VERSION : 1.2
// clk_pulse uses the internal sps time to generate a clock with programmable period time.
// the period time is defined for 10ms .. 65s.
// pulse generation is continuous if N = 0 and for n pulses otherwise.
// the first cycle after start is a clk pulse and then depending on the programmed period time a delay.
// every pulse is only valid for one cycle so that a edge trigger is not necessary
// clk_prg depending on the accuracy of the system clock.
// 
// uses: T_PLC_MS [FC64]
//       STIME [FB64],IDB_STIME [DB64]
   VAR_INPUT
      PT : Time;
      N : Int;
      RST : Bool;
   END_VAR
   VAR_OUTPUT
      Q : Bool;
      CNT : Int;
      RUN : Bool;
   END_VAR
   VAR
      tx : DWord;
      tn : DWord;
      init : Bool;
   END_VAR
   VAR_TEMP
      TOP_SI : Struct
         EV_CLASS : Byte;
         EV_NUM : Byte;
         PRIORITY : Byte;
         NUM : Byte;
         TYP2_3 : Byte;
         TYP1 : Byte;
         ZI1 : Word;
         ZI2_3 : DWord;
      END_STRUCT;
      START_UP_SI : Struct
         EV_CLASS : Byte;
         EV_NUM : Byte;
         PRIORITY : Byte;
         NUM : Byte;
         TYP2_3 : Byte;
         TYP1 : Byte;
         ZI1 : Word;
         ZI2_3 : DWord;
      END_STRUCT;
      ERR : Int;
   END_VAR
BEGIN


   (* read actual startup info *)
   (* OB1_SCAN_1  BYTE  -  B#16#01: Abschluss des Neustarts (Warmstarts)
                        -  B#16#02: Abschluss des Wiederanlaufs
                        -  B#16#03: Abschluss des freien Zyklus
                        -  B#16#04: Abschluss des Kaltstarts
                        -  B#16#05: Erster OB 1-Zyklus der neuen Master-CPU nach 
                                    Master-Reserve-Umschaltung und STOP des 
                                    bisherigen Masters *)

     #ERR := RD_SINFO (TOP_SI => #TOP_SI, START_UP_SI => #START_UP_SI);

   (* detect system startup *)
     IF #TOP_SI.EV_NUM = 1 OR #TOP_SI.EV_NUM = 2 OR #TOP_SI.EV_NUM = 4 THEN 
       #init := FALSE;
     END_IF;

     #tx := "T_PLC_MS"();   (* read system *)
     #Q := FALSE;       (* reset Q we generate pulses only for one cycle *)
     #RUN := #CNT < #N;

     IF NOT #init OR #RST THEN
       #init := TRUE;
       #CNT := 0;
       #tn := DINT_TO_DWORD(DWORD_TO_DINT(#tx) - T_CONV(#PT));
       #RUN := FALSE;
     ELSIF (#CNT < #N OR #N = 0) AND DWORD_TO_DINT(#tx) - DWORD_TO_DINT(#tn) >= T_CONV(#PT) THEN    (* generate a pulse *)
       #CNT := #CNT + 1;
       #Q := TRUE;
       #tn := DINT_TO_DWORD(DWORD_TO_DINT(#tn) + T_CONV(#PT));
     END_IF;


   (* revision history
   hm    4. aug 2006   rev 1.0
     original version

   hm    17. sep 2007  rev 1.1
     replaced time() with T_PLC_S() for compatblity reasons

   hm    16. feb. 2011 rev 1.2
     fixed an error when timer overflows 
   *)
END_FUNCTION_BLOCK

FUNCTION_BLOCK "D_TRIG"   // FB54, SCL
TITLE = D_TRIG
{ S7_Optimized_Access := 'FALSE' }
AUTHOR : hugo
FAMILY : GENERAT
NAME : D_TRIG
VERSION : 1.1
// this block is similar to the IEC Standard R_trig and F_trig but it monitors a DWORD, WORD or Byte Variable instead and generated an Output Pulse for one cycle only when the input has changed.
// an additional output x (Dword) will state the chage of the input.
// Example: the input has chaged from 0001 to 0010 then the output x will be 2.
   VAR_INPUT
      in : DWord;
   END_VAR
   VAR_OUTPUT
      Q : Bool;
      X : DWord;
   END_VAR
   VAR
      last_in : DWord;
   END_VAR
BEGIN


     #Q := #in <> #last_in;
     #X := DINT_TO_DWORD(DWORD_TO_DINT(#in) - DWORD_TO_DINT(#last_in));
     #last_in := #in;


   (* revision history

   hm  4.09.2007   rev 1.0
     original version released

   hm  19. feb. 2008 rev 1.1
     performance improvement
   *)
END_FUNCTION_BLOCK

FUNCTION_BLOCK "GEN_BIT"   // FB55, SCL
TITLE = GEN_BIT
{ S7_Optimized_Access := 'FALSE' }
AUTHOR : hugo
FAMILY : GENERAT
NAME : GEN_BIT
VERSION : 1.2
// gen_bit is 4 bit sequencial pattern generator with 4 DWORD inputs and 4 serial outputs.
// with the first clock pulse after a reset or after power on, bit 0 of the input DWORDS IN is present on the Outputs Q and the next clock cycle shifts to Bit 1 and so on.
// the input steps defines how many bits of the input dwords will be shifted to the outputs. the sequence can be repetive when rep = 0 or any amount of repetitions can be defined with input rep.
   VAR_INPUT
      in0 : DWord;
      in1 : DWord;
      in2 : DWord;
      in3 : DWord;
      clk : Bool;
      steps : Int;
      rep : Int;
      rst : Bool;
   END_VAR
   VAR_OUTPUT
      Q0 : Bool;
      Q1 : Bool;
      Q2 : Bool;
      Q3 : Bool;
      cnt : Int;
      run : Bool;
   END_VAR
   VAR
      r0 : DWord;
      tr0 AT r0 : Array[0..31] of Bool;
      r1 : DWord;
      tr1 AT r1 : Array[0..31] of Bool;
      r2 : DWord;
      tr2 AT r2 : Array[0..31] of Bool;
      r3 : DWord;
      tr3 AT r3 : Array[0..31] of Bool;
      rx : Int := 1;
   END_VAR
BEGIN


   (* check if number of runs is finished or rep = 0 which means continuous *)
   IF #clk AND NOT #rst THEN
       #run := (#rep = 0) OR (#rx <= #rep);
       IF #run THEN
           (* check for step counter reached and reset to 0 if cnt = steps *)
           IF #cnt = #steps THEN
               #cnt := 0;
           END_IF;

           (* when cnt = 0 then reload the inputs into the registers *)
           IF #cnt = 0 THEN
               #r0 := #in0;
               #r1 := #in1;
               #r2 := #in2;
               #r3 := #in3;
           END_IF;

           (* when cnt < steps, shift the lowest bits to the outputs *)
           IF (#cnt < #steps) THEN
               #Q0 := #tr0[24];
               #Q1 := #tr1[24];
               #Q2 := #tr2[24];
               #Q3 := #tr3[24];
               #r0 := SHR(IN:=#r0,N:=1);
               #r1 := SHR(IN:=#r1,N:=1);
               #r2 := SHR(IN:=#r2,N:=1);
               #r3 := SHR(IN:=#r3,N:=1);
           END_IF;

           (* increment the step counter *)
           #cnt := #cnt +1;
           IF (#cnt = #steps) AND (#rep <> 0) THEN #rx := #rx +1; END_IF;
           IF (#rx > #rep) AND (#rep <> 0) THEN #run := FALSE; END_IF;
       END_IF;
   ELSE
       IF #rst THEN
           #run := FALSE;
           #Q0 := FALSE;
           #Q1 := FALSE;
           #Q2 := FALSE;
           #Q3 := FALSE;
           #r0 := 0;
           #r1 := 0;
           #r2 := 0;
           #r3 := 0;
           #cnt := 0;
           #rx := 1;
       END_IF;
   END_IF;


   (* revision histroy
   hm  4 aug 2006  rev 1.0
       original version

   hm 15. oct. 2008    rev 1.1
       improved performance

   hm  14. mar. 2009   rev 1.2
       removed double assignments

   *)
END_FUNCTION_BLOCK

FUNCTION_BLOCK "GEN_SQ"   // FB56, SCL
TITLE = GEN_SQ
{ S7_Optimized_Access := 'FALSE' }
AUTHOR : hugo
FAMILY : GENERAT
NAME : GEN_SQ
VERSION : 1.3
// gen_sq generates square wave signal with programmable period time.
// 
// uses: T_PLC_MS [FC64]
//       STIME [FB64],IDB_STIME [DB64]
   VAR_INPUT
      PT : Time;
   END_VAR
   VAR_OUTPUT
      Q : Bool;
   END_VAR
   VAR
      tn : Time;
      tx : Time;
      init : Bool;
   END_VAR
   VAR_TEMP
      TOP_SI : Struct
         EV_CLASS : Byte;
         EV_NUM : Byte;
         PRIORITY : Byte;
         NUM : Byte;
         TYP2_3 : Byte;
         TYP1 : Byte;
         ZI1 : Word;
         ZI2_3 : DWord;
      END_STRUCT;
      START_UP_SI : Struct
         EV_CLASS : Byte;
         EV_NUM : Byte;
         PRIORITY : Byte;
         NUM : Byte;
         TYP2_3 : Byte;
         TYP1 : Byte;
         ZI1 : Word;
         ZI2_3 : DWord;
      END_STRUCT;
      ERR : Int;
   END_VAR
BEGIN


     (* read actual startup info *)
     (* OB1_SCAN_1  BYTE  -  B#16#01: Abschluss des Neustarts (Warmstarts)
                          -  B#16#02: Abschluss des Wiederanlaufs
                          -  B#16#03: Abschluss des freien Zyklus
                          -  B#16#04: Abschluss des Kaltstarts
                          -  B#16#05: Erster OB 1-Zyklus der neuen Master-CPU nach 
                                      Master-Reserve-Umschaltung und STOP des 
                                      bisherigen Masters *)

     #ERR := RD_SINFO (TOP_SI => #TOP_SI, START_UP_SI => #START_UP_SI);

     (* read system time *)
     #tx := T_CONV(DWORD_TO_DINT("T_PLC_MS"()));

     (* reset last_time on system startup *)
     IF #TOP_SI.EV_NUM = 1 OR #TOP_SI.EV_NUM = 2 OR #TOP_SI.EV_NUM = 4 THEN 
       #init := FALSE;
     END_IF;

     IF NOT #init THEN
       #init := TRUE;
       #tn := #tx;
       #Q := TRUE;
     ELSIF #tx - #tn >= T_CONV(DWORD_TO_DINT(SHR(IN:=DINT_TO_DWORD(T_CONV(#PT)),N:=1))) THEN
       #Q := NOT #Q;
       #tn := #tn + T_CONV(DWORD_TO_DINT(SHR(IN:=DINT_TO_DWORD(T_CONV(#PT)),N:=1)));
     END_IF;


   (* revision history
   hm  4. aug 2006 rev 1.0
     original version

   hm  17. sep 2007  rev 1.1
     replaced time() with T_PLC_MS() for compatibility reasons

   hm  18. jul. 2009 rev 1.2
     improved accuracy

   hm  16. feb 2011  rev 1.3
     corrected an error with timer overflow 
   *)
END_FUNCTION_BLOCK

FUNCTION_BLOCK "SCHEDULER"   // FB57, SCL
TITLE = SCHEDULER
{ S7_Optimized_Access := 'FALSE' }
AUTHOR : hugo
FAMILY : GENERAT
NAME : SCHED
VERSION : 1.1
// SCHEDULER is used to call programs or function blocks at specific intervals.
// T0..T3 defines the interval times.
// 
// uses: T_PLC_MS [FC64]
//       STIME [FB64],IDB_STIME [DB64]
   VAR_INPUT
      E0 : Bool;
      E1 : Bool;
      E2 : Bool;
      E3 : Bool;
      T_0 : Time;
      T_1 : Time;
      T_2 : Time;
      T_3 : Time;
   END_VAR
   VAR_OUTPUT
      Q0 : Bool;
      Q1 : Bool;
      Q2 : Bool;
      Q3 : Bool;
   END_VAR
   VAR
      init : Bool;
      s0 : Time;
      s1 : Time;
      s2 : Time;
      s3 : Time;
      tx : Time;
      c : Int;
   END_VAR
BEGIN


   (* read system_time *)
   #tx := T_CONV(DWORD_TO_DINT("T_PLC_MS"()));

   IF NOT #init THEN
       #init := TRUE;
       #s0 := #tx - #T_0;
       #s1 := #tx - #T_1;
       #s2 := #tx - #T_2;
       #s3 := #tx - #T_3;
   END_IF;

   #Q0 := FALSE;
   #Q1 := FALSE;
   #Q2 := FALSE;
   #Q3 := FALSE;

   CASE #c OF
       0:  IF #tx - #s0 >= #T_0 THEN
               #Q0 := #E0;
               #s0 := #tx;
           END_IF;
           #c := 1;
       1:  IF #tx - #s1 >= #T_1 THEN
               #Q1 := #E1;
               #s1 := #tx;
           END_IF;
           #c := 2;
       2:  IF #tx - #s2 >= #T_2 THEN
               #Q2 := #E2;
               #s2 := #tx;
           END_IF;
           #c := 3;
       3:  IF #tx - #s3 >= #T_3 THEN
               #Q3 := #E3;
               #s3 := #tx;
           END_IF;
           #c := 0;
   END_CASE;


   (* revision history

   hm 28. sep. 2008    rev 1.0
       original version

   hm  14. mar. 2009   rev 1.1
       removed double assignments

   *)
END_FUNCTION_BLOCK

FUNCTION_BLOCK "SCHEDULER_2"   // FB58, SCL
TITLE = SCHEDULER_2
{ S7_Optimized_Access := 'FALSE' }
AUTHOR : hugo
FAMILY : GENERAT
NAME : SCHED2
VERSION : 1.0
// SCHEDULER_2 is used to call programs or function blocks at specific cycles.
// C0..C3 defines after how many cycles the output becomes active.
// O0..O3 defines a cycle offset at startup.
   VAR_INPUT
      E0 : Bool;
      E1 : Bool;
      E2 : Bool;
      E3 : Bool;
      C0 : Int;
      C1 : Int;
      C2 : Int;
      C3 : Int;
      O0 : Int;
      O1 : Int;
      O2 : Int;
      O3 : Int;
   END_VAR
   VAR_OUTPUT
      Q0 : Bool;
      Q1 : Bool;
      Q2 : Bool;
      Q3 : Bool;
   END_VAR
   VAR
      sx : Int;
   END_VAR
BEGIN


   #Q0 := #E0 AND (#sx MOD #C0 - #O0 = 0);
   #Q1 := #E1 AND (#sx MOD #C1 - #O1 = 0);
   #Q2 := #E2 AND (#sx MOD #C2 - #O2 = 0);
   #Q3 := #E3 AND (#sx MOD #C3 - #O3 = 0);

   (* increment cycle counter every cycle *)
   #sx := #sx + 1;


   (* revision history
   hm 29. sep. 2008        rev 1.0
       original version


   *)
END_FUNCTION_BLOCK

FUNCTION_BLOCK "SEQUENCE_4"   // FB59, SCL
TITLE = SEQUENCE_4
{ S7_Optimized_Access := 'FALSE' }
AUTHOR : oscat
FAMILY : GENERAT
NAME : SEQ_4
VERSION : 1.5
// sequence_4 enables run when a low to high transition is present on start.
// a low to high transition on start will restart the sequencer at any time while a rst will hold the sequencer in reset while true.
// after run is enabled with a rising edge on start the sequencer waits for wait0 on in0 to enable q0 which stays on for delay0.
// the next cycle starts with wait1, continues with delay 1 and so on...
// if an edge is not detected during the wait period, the sequencer will then display the error number on the status output.
// the status numbers 1..4 are errors in step 0..3.
// after the last step that sets q3, the sequencer leaves q3 on for delay3 and then resets to the initial state.
// a step output will indicate the current step of the sequencer and will also be present with a fault condition.
// after the first output is turened on the sequencer switches from q0 to q1 and so on, at any time there is only one output enabled.
// if an input signal is not detected during a wait period, the sequencer will display the error number ( 1 for in0, 2 for in1 .... ).
// when an error is present and the config variable stop_on_error is set then the sequencer will stop. otherwise it will continue.
// The status output will also display 110 for waiting and 111 for sequence running.
// 
// uses: T_PLC_MS [FC64]
//       STIME [FB64],IDB_STIME [DB64]
   VAR_INPUT
      in0 : Bool := TRUE;
      in1 : Bool := TRUE;
      in2 : Bool := TRUE;
      in3 : Bool := TRUE;
      start : Bool;
      rst : Bool;
      wait0 : Time;
      delay0 : Time;
      wait1 : Time;
      delay1 : Time;
      wait2 : Time;
      delay2 : Time;
      wait3 : Time;
      delay3 : Time;
      stop_on_error : Bool;
   END_VAR
   VAR_OUTPUT
      Q0 : Bool;
      Q1 : Bool;
      Q2 : Bool;
      Q3 : Bool;
      QX : Bool;
      run : Bool;
      "step" : Int := -1;
      status : Byte;
   END_VAR
   VAR
      last : Time;
      edge : Bool;
      tx : Time;
      init : Bool;
   END_VAR
BEGIN


   (* read sps timer *)
   #tx := T_CONV(DWORD_TO_DINT("T_PLC_MS"()));

   (* initialize on startup *)
   IF NOT #init THEN
       #last := #tx;
       #init := TRUE;
       #status := 110;
   END_IF;

   (* asynchronous reset *)
   IF #rst THEN
       #"step" := -1;
       #Q0 := 0;
       #Q1 := 0;
       #Q2 := 0;
       #Q3 := 0;
       #status := 110;
       #run := 0;

     (* edge on start input restarts the sequencer *)
   ELSIF #start AND NOT #edge THEN
       #"step" := 0;
       #last := #tx;
       #status := 111;
       #Q0 := 0;
       #Q1 := 0;
       #Q2 := 0;
       #Q3 := 0;
       #run := 1;
   END_IF;
   #edge := #start;

   (* check if stop on status is necessary *)
   IF BYTE_TO_INT(#status) > 0 AND BYTE_TO_INT(#status) < 100 AND #stop_on_error THEN RETURN; END_IF;

   (* sequence is running *)
   IF #run AND #"step" = 0 THEN
       IF NOT #Q0 AND #in0 AND #tx - #last <= #wait0 THEN
           #Q0 := TRUE;
           #last := #tx;
       ELSIF NOT #Q0 AND #tx - #last > #wait0 THEN
           #status := 1;
           #run := FALSE;
       ELSIF #Q0 AND #tx - #last >= #delay0 THEN
           #"step" := 1;
           #last := #tx;
       END_IF;
   END_IF;
   IF #run AND #"step" = 1 THEN
       IF NOT #Q1 AND #in1 AND #tx - #last <= #wait1 THEN
         #Q0 := FALSE;
         #Q1 := TRUE;
         #last := #tx;
       ELSIF NOT #Q1 AND #tx - #last > #wait1 THEN
         #status := 2;
         #Q0 := FALSE;
         #run := FALSE;
       ELSIF #Q1 AND #tx - #last >= #delay1 THEN
         #"step" := 2;
         #last := #tx;
       END_IF;
   END_IF;
   IF #run AND #"step" = 2 THEN
       IF NOT #Q2 AND #in2 AND #tx - #last <= #wait2 THEN
         #Q1 := FALSE;
         #Q2 := TRUE;
         #last := #tx;
       ELSIF NOT #Q2 AND #tx - #last > #wait2 THEN
         #status := 3;
         #Q1 := FALSE;
         #run := FALSE;
       ELSIF #Q2 AND #tx - #last >= #delay2 THEN
         #"step" := 3;
         #last := #tx;
       END_IF;
   END_IF;
   IF #run AND #"step" = 3 THEN
       IF NOT #Q3 AND #in3 AND #tx - #last <= #wait3 THEN
         #Q2 := FALSE;
         #Q3 := TRUE;
         #last := #tx;
       ELSIF NOT #Q3 AND #tx - #last > #wait3 THEN
         #status := 4;
         #Q2 := FALSE;
         #run := FALSE;
       ELSIF #Q3 AND #tx - #last >= #delay3 THEN
         #"step" := -1;
         #Q3 := FALSE;
         #run := FALSE;
         #status := 110;
       END_IF;
   END_IF;
   #QX := #Q0 OR #Q1 OR #Q2 OR #Q3;


   (*
   hm 1.10.06      rev 1.1
       corrected delay logic to be after event and not before
       added any output

   hm 1.12.06      rev 1.2
       corrected failure in sequence logic.
       added init at startup to prevent from initial error after start.

   hm 17.1.2007        rev 1.3
       changed output fault to status for better compatibility with other modules (ESR).
       added stop on error functionality and setup variable
       default for inputs in0..3 is true.
       renamed variable state to step

   hm  17.sep 2007 rev 1.4
       replaced time() with T_PLC_MS() for compatibility reasons

   hm  13. mar. 2009   rev 1.5
       renamed output any to qx for compatibility resons

   *)
END_FUNCTION_BLOCK

FUNCTION_BLOCK "SEQUENCE_64"   // FB60, SCL
TITLE = SEQUENCE_64
{ S7_Optimized_Access := 'FALSE' }
AUTHOR : hugo
FAMILY : GENERAT
NAME : SEQ_64
VERSION : 1.0
// sequence generates a sequence of states with a programmable length for each state.
// 
// uses: T_PLC_MS [FC64]
//       STIME [FB64],IDB_STIME [DB64]
//       INC2 [FC91]
   VAR_INPUT
      START : Bool;
      SMAX : Int;
      PROG : Array[0..63] of Time;
      RST : Bool;
   END_VAR
   VAR_OUTPUT
      STATE : Int := -1;
      TRIG : Bool;
   END_VAR
   VAR
      tx : Time;
      edge : Bool;
      last : Time;
   END_VAR
BEGIN


   (* read system timer *)
   #tx := T_CONV(DWORD_TO_DINT("T_PLC_MS"()));
   #TRIG := FALSE;

   IF #RST THEN
       #STATE := -1;

   (* start sequence *)
   ELSIF #START AND NOT #edge THEN
       #STATE := 0;
       #last := #tx;
       #TRIG := TRUE;

   (* sequence generator *)
   ELSIF (#STATE >= 0) THEN
       IF (#tx - #last) >= #PROG[#STATE] THEN
           #STATE := "INC2"(X:=#STATE,D:=1,L:=-1,U:=#SMAX);
           #last := #tx;
           #TRIG := TRUE;
       END_IF;
   END_IF;

   #edge := #START;



   (* revision history
   hm  29. jun. 2008
       original version

   *)
END_FUNCTION_BLOCK

FUNCTION_BLOCK "SEQUENCE_8"   // FB61, SCL
TITLE = SEQUENCE_8
{ S7_Optimized_Access := 'FALSE' }
AUTHOR : oscat
FAMILY : GENERAT
NAME : SEQ_8
VERSION : 1.5
// sequence_8 enables run when a low to high transition is present on start.
// a low to high transition on start will restart the sequencer at any time while a rst will hold the sequencer in reset while true.
// after run is enabled with a rising edge on start the sequencer waits for wait0 on in0 to enable q0 which stays on for delay0.
// the next cycle starts with wait1, continues with delay 1 and so on...
// if an edge is not detected during the wait period, the sequencer will then display the error number on the status output.
// The status numbers are 1 .. 8 for erros in step 0..7.
// after the last step that sets q7, the sequencer leaves q7 on for delay7 and then resets to the initial state.
// a step output will indicate the current step of the sequencer and will also be present with a fault condition.
// after the first output is turened on the sequencer switches from q0 to q1 and so on, at any time there is only one output enabled.
// if an input signal is not detected during a wait period, the sequencer will display the error number ( 1 for in0, 2 for in1 .... ).
// when an error is present and the config variable stop_on_error is set then the sequencer will stop. otherwise it will continue.
// The status output will also display 110 for waiting and 111 sequece running.
// 
// uses: T_PLC_MS [FC64]
//       STIME [FB64],IDB_STIME [DB64]
   VAR_INPUT
      in0 : Bool := TRUE;
      in1 : Bool := TRUE;
      in2 : Bool := TRUE;
      in3 : Bool := TRUE;
      in4 : Bool := TRUE;
      in5 : Bool := TRUE;
      in6 : Bool := TRUE;
      in7 : Bool := TRUE;
      start : Bool;
      rst : Bool;
      wait0 : Time;
      delay0 : Time;
      wait1 : Time;
      delay1 : Time;
      wait2 : Time;
      delay2 : Time;
      wait3 : Time;
      delay3 : Time;
      wait4 : Time;
      delay4 : Time;
      wait5 : Time;
      delay5 : Time;
      wait6 : Time;
      delay6 : Time;
      wait7 : Time;
      delay7 : Time;
      stop_on_error : Bool;
   END_VAR
   VAR_OUTPUT
      Q0 : Bool;
      Q1 : Bool;
      Q2 : Bool;
      Q3 : Bool;
      Q4 : Bool;
      Q5 : Bool;
      Q6 : Bool;
      Q7 : Bool;
      QX : Bool;
      run : Bool;
      "step" : Int := -1;
      status : Byte;
   END_VAR
   VAR
      last : Time;
      edge : Bool;
      tx : Time;
      init : Bool;
   END_VAR
BEGIN


   (* read sps timer *)
   #tx := T_CONV(DWORD_TO_DINT("T_PLC_MS"()));

   (* initialize on startup *)
   IF NOT #init THEN
       #last := #tx;
       #init := TRUE;
       #status := 110;
   END_IF;

   (* asynchronous reset *)
   IF #rst THEN
       #"step" := -1;
       #Q0 := 0;
       #Q1 := 0;
       #Q2 := 0;
       #Q3 := 0;
       #Q4 := 0;
       #Q5 := 0;
       #Q6 := 0;
       #Q7 := 0;
       #status := 110;
       #run := 0;

   (* edge on start input restarts the sequencer *)
   ELSIF #start AND NOT #edge THEN
       #"step" := 0;
       #last := #tx;
       #status := 111;
       #Q0 := 0;
       #Q1 := 0;
       #Q2 := 0;
       #Q3 := 0;
       #Q4 := 0;
       #Q5 := 0;
       #Q6 := 0;
       #Q7 := 0;
       #run := 1;
     END_IF;
     #edge := #start;

   (* check if stop on error is necessary *)
   IF BYTE_TO_INT(#status) > 0 AND BYTE_TO_INT(#status) < 100 AND #stop_on_error THEN RETURN; END_IF;

   (* sequence is running *)
   IF #run AND #"step" = 0 THEN
       IF NOT #Q0 AND #in0 AND #tx - #last <= #wait0 THEN
           #Q0 := TRUE;
           #last := #tx;
       ELSIF NOT #Q0 AND #tx - #last > #wait0 THEN
           #status := 1;
           #run := FALSE;
       ELSIF #Q0 AND #tx - #last >= #delay0 THEN
           #"step" := 1;
           #last := #tx;
       END_IF;
   END_IF;
   IF #run AND #"step" = 1 THEN
       IF NOT #Q1 AND #in1 AND #tx - #last <= #wait1 THEN
           #Q0 := FALSE;
           #Q1 := TRUE;
           #last := #tx;
       ELSIF NOT #Q1 AND #tx - #last > #wait1 THEN
           #status := 2;
           #Q0 := FALSE;
           #run := FALSE;
       ELSIF #Q1 AND #tx - #last >= #delay1 THEN
           #"step" := 2;
           #last := #tx;
       END_IF;
   END_IF;
   IF #run AND #"step" = 2 THEN
       IF NOT #Q2 AND #in2 AND #tx - #last <= #wait2 THEN
           #Q1 := FALSE;
           #Q2 := TRUE;
           #last := #tx;
       ELSIF NOT #Q2 AND #tx - #last > #wait2 THEN
           #status := 3;
           #Q1 := FALSE;
           #run := FALSE;
       ELSIF #Q2 AND #tx - #last >= #delay2 THEN
           #"step" := 3;
           #last := #tx;
       END_IF;
   END_IF;
   IF #run AND #"step" = 3 THEN
       IF NOT #Q3 AND #in3 AND #tx - #last <= #wait3 THEN
           #Q2 := FALSE;
           #Q3 := TRUE;
           #last := #tx;
       ELSIF NOT #Q3 AND #tx - #last > #wait3 THEN
           #status := 4;
           #Q2 := FALSE;
           #run := FALSE;
       ELSIF #Q3 AND #tx - #last >= #delay3 THEN
           #"step" := 4;
           #last := #tx;
       END_IF;
   END_IF;
   IF #run AND #"step" = 4 THEN
       IF NOT #Q4 AND #in4 AND #tx - #last <= #wait4 THEN
           #Q3 := FALSE;
           #Q4 := TRUE;
           #last := #tx;
       ELSIF NOT #Q4 AND #tx - #last > #wait4 THEN
           #status := 5;
           #Q3 := FALSE;
           #run := FALSE;
       ELSIF #Q4 AND #tx - #last >= #delay4 THEN
           #"step" := 5;
           #last := #tx;
       END_IF;
   END_IF;
   IF #run AND #"step" = 5 THEN
       IF NOT #Q5 AND #in5 AND #tx - #last <= #wait5 THEN
           #Q4 := FALSE;
           #Q5 := TRUE;
           #last := #tx;
       ELSIF NOT #Q5 AND #tx - #last > #wait5 THEN
           #status := 6;
           #Q4 := FALSE;
           #run := FALSE;
       ELSIF #Q5 AND #tx - #last >= #delay5 THEN
           #"step" := 6;
           #last := #tx;
       END_IF;
   END_IF;
   IF #run AND #"step" = 6 THEN
       IF NOT #Q6 AND #in6 AND #tx - #last <= #wait6 THEN
           #Q5 := FALSE;
           #Q6 := TRUE;
           #last := #tx;
       ELSIF NOT #Q6 AND #tx - #last > #wait6 THEN
           #status := 7;
           #Q5 := FALSE;
           #run := FALSE;
       ELSIF #Q6 AND #tx - #last >= #delay6 THEN
           #"step" := 7;
           #last := #tx;
       END_IF;
   END_IF;
   IF #run AND #"step" = 7 THEN
       IF NOT #Q7 AND #in7 AND #tx - #last <= #wait7 THEN
           #Q6 := FALSE;
           #Q7 := TRUE;
           #last := #tx;
       ELSIF NOT #Q7 AND #tx - #last > #wait7 THEN
           #status := 8;
           #Q6 := FALSE;
           #run := FALSE;
       ELSIF #Q7 AND #tx - #last >= #delay7 THEN
           #"step" := -1;
           #Q7 := FALSE;
           #run := FALSE;
           #status := 110;
       END_IF;
   END_IF;
   #QX := #Q0 OR #Q1 OR #Q2 OR #Q3 OR #Q4 OR #Q5 OR #Q6 OR #Q7;


   (*
   hm 1.10.06      rev 1.1
       corrected delay logic to be after event and not before
       added any output

   hm 1.12.06      rev 1.2
       corrected failure in sequence logic.
       added init at startup to prevent from initial statuss after start.

   hm 17.1.2007        rev 1.3
       changed output fault to status for better compatibility with other modules (ESR)
       added stop on error functionality and setup variable
       default for inputs in0..7 is true.
       renames variable state to step

   hm  17.sep 2007 rev 1.4
       replaced time() with T_PLC_MS() for compatibility reasons

   hm  13. mar. 2009   rev 1.5
       renamed output any to qx for compatibility resons

   *)
END_FUNCTION_BLOCK

FUNCTION_BLOCK "TMAX"   // FB62, SCL
TITLE = TMAX
{ S7_Optimized_Access := 'FALSE' }
AUTHOR : hugo
FAMILY : GENERAT
NAME : TMAX
VERSION : 1.0
// Q of tmax will follow IN except that it forces a maximum ontime for the output Q.
// the output Z will be active for one cycle if the output is forced low by the timeout.
// 
// uses: T_PLC_MS [FC64]
//       STIME [FB64],IDB_STIME [DB64]
   VAR_INPUT
      IN : Bool;
      PT : Time;
   END_VAR
   VAR_OUTPUT
      Q : Bool;
      Z : Bool;
   END_VAR
   VAR
      tx : Time;
      start : Time;
      last_in : Bool;
   END_VAR
BEGIN


   (* read system timer *)
   #tx := T_CONV(DWORD_TO_DINT("T_PLC_MS"()));

   #Z := FALSE;

   IF NOT #IN THEN
       #Q := FALSE;
   ELSIF #IN AND NOT #last_in THEN
       #Q := TRUE;
       #start := #tx;
   ELSIF (#tx - #start >= #PT) AND #Q THEN
       #Q := FALSE;
       #Z := TRUE;
   END_IF;

   #last_in := #IN;



   (* revision history
   hm  20. jul. 2008   rev 1.0
       original version

   *)
END_FUNCTION_BLOCK

FUNCTION_BLOCK "TMIN"   // FB63, SCL
TITLE = TMIN
{ S7_Optimized_Access := 'FALSE' }
AUTHOR : hugo
FAMILY : GENERAT
NAME : TMIN
VERSION : 1.0
// Q of tMIN will follow IN except that it forces a minimum ontime for the output Q.
   VAR_INPUT
      IN : Bool;
      PT : Time;
   END_VAR
   VAR_OUTPUT
      Q : Bool;
   END_VAR
   VAR
      pm : TP;
   END_VAR
BEGIN


   #pm(IN := #IN, PT := #PT);
   #Q := #IN OR #pm.Q;


   (* revision history
   hm  21. jul. 2008   rev 1.0
       original version

   *)
END_FUNCTION_BLOCK

FUNCTION_BLOCK "STIME"   // FB64, SCL
TITLE = STIME
{ S7_Optimized_Access := 'FALSE' }
AUTHOR : dalbi
FAMILY : MEASURE
NAME : STIME
VERSION : 1.4
// this function block makes sure that the timer of a siemens sps counts from 0 - 2^32-1.
   VAR_OUTPUT
      tx : DWord;
      at_tx AT tx : Array[0..31] of Bool;
   END_VAR
   VAR
      last_time : DWord;
      bit31 : Bool;
      init : Bool := TRUE;
   END_VAR
   VAR_TEMP
      TOP_SI : Struct
         EV_CLASS : Byte;
         EV_NUM : Byte;
         PRIORITY : Byte;
         NUM : Byte;
         TYP2_3 : Byte;
         TYP1 : Byte;
         ZI1 : Word;
         ZI2_3 : DWord;
      END_STRUCT;
      START_UP_SI : Struct
         EV_CLASS : Byte;
         EV_NUM : Byte;
         PRIORITY : Byte;
         NUM : Byte;
         TYP2_3 : Byte;
         TYP1 : Byte;
         ZI1 : Word;
         ZI2_3 : DWord;
      END_STRUCT;
      ERR : Int;
   END_VAR
BEGIN


   (* this FB is only necessary for siemens sps
   the siemens sps timer counts from 0 to 2^31-1 and starts at 0 sfter overrun.
   this means that the bit 31 (the highest bit ) will never be used and therefore
   a problem arises when t2 - t1 is checked.
   t2 - t1 is always valid also in an timer overrun situation where the time t1 is very high and t2 is very low.
   the result of the subtraction t2 - t1 however is still valid.
   this calculation does not work for soiemens because the highest bit is not used.

   this module stores the highest bit, changes the highest bit at every overrun occurence and stuffs ther highest bit in the output.
   the output is then used by t_plc_us and t_plc_ms.

   the correction needs and fb and not a function because the value of the highest bit has to be stored.

   do never use this function block in a codesys environment. the timer in codesys is correct and runs from 0 to 2^32-1
   *)

   (* read actual startup info *)
   (* OB1_SCAN_1  BYTE  -  B#16#01: Abschluss des Neustarts (Warmstarts)
                        -  B#16#02: Abschluss des Wiederanlaufs
                        -  B#16#03: Abschluss des freien Zyklus
                        -  B#16#04: Abschluss des Kaltstarts
                        -  B#16#05: Erster OB 1-Zyklus der neuen Master-CPU nach 
                                    Master-Reserve-Umschaltung und STOP des 
                                    bisherigen Masters *)

   #ERR := RD_SINFO (TOP_SI => #TOP_SI, START_UP_SI => #START_UP_SI);

   (* reset last_time on system startup *)
   IF #TOP_SI.EV_NUM = 1 OR #TOP_SI.EV_NUM = 2 OR #TOP_SI.EV_NUM = 4 OR NOT #init THEN 
       #last_time := 0;
       #bit31 := false;
       #init := true;
   END_IF;

   (* read the system timer *)
   #tx := DINT_TO_DWORD(T_CONV(TIME_TCK()));

   (* check for overrun *)
   IF DWORD_TO_DINT(#tx) < DWORD_TO_DINT(#last_time) THEN
       (* an overrun has occured, change the value of the highest bit *)
       #bit31 := NOT #bit31;
   END_IF;

   (* stuff the highest bit into the timer value *)
   #at_tx[7] := #bit31;

   (* remember the last system time for the next overrun check *)
   #last_time := #tx;


   (* revision history
   DA  14.9.2007 rev 1.0
     original version

   DA  24.2.2008 rev 1.1
     added self reset on system startup

   DA   2.5.2008 rev 1.2
     corect a problem running under OB35

   DA  12.3.2009 rev 1.3
     corect a problem run on different CPUs

   DA  22.12.2009 rev 1.4
     corect a problem on startup
   *)
END_FUNCTION_BLOCK

FUNCTION_BLOCK "TOF_1"   // FB65, SCL
TITLE = TOF_1
{ S7_Optimized_Access := 'FALSE' }
AUTHOR : hugo
FAMILY : GENERAT
NAME : TOF_1
VERSION : 1.0
// TOF_1 will extend a pulse on input in for PT seconds.
// in addition the timer can be cleared asynchronously with rst.
// TOF_1 is the same function as TOF from the standard LIB except the asynchronous reset input.
// 
// uses: T_PLC_MS [FC64]
//       STIME [FB64],IDB_STIME [DB64]
   VAR_INPUT
      IN : Bool;
      PT : Time;
      RST : Bool;
   END_VAR
   VAR_OUTPUT
      Q : Bool;
   END_VAR
   VAR
      tx : Time;
      start : Time;
   END_VAR
BEGIN


   (* read system timer *)
   #tx := T_CONV(DWORD_TO_DINT("T_PLC_MS"()));

   IF #RST THEN
       #Q := FALSE;
   ELSIF #IN THEN
       #Q := TRUE;
       #start := #tx;
   ELSIF #tx - #start >= #PT THEN
       #Q := FALSE;
   END_IF;




   (* revision history
   hm  17. jul. 2008   rev 1.0
       original version

   *)
END_FUNCTION_BLOCK

FUNCTION_BLOCK "TONOF"   // FB66, SCL
TITLE = TONOF
{ S7_Optimized_Access := 'FALSE' }
AUTHOR : hugo
FAMILY : GENERAT
NAME : TONOF
VERSION : 1.2
// TONOF generated a TON and TOF Delay for the Input N TON (T1) and TOF (T2) can be configured separately
   VAR_INPUT
      IN : Bool;
      T_ON : Time;
      T_OFF : Time;
   END_VAR
   VAR_OUTPUT
      Q : Bool;
   END_VAR
   VAR
      X : TON;
      old : Bool;
      mode : Bool;
   END_VAR
BEGIN


   IF #IN XOR #old THEN
     #X(IN := FALSE, PT := SEL(G := #IN, IN0 := #T_OFF, IN1 := #T_ON));
     #mode := #IN;
     #old := #IN;
   END_IF;
   #X.IN := TRUE;
   IF #X.Q THEN #Q := #mode;END_IF;


   (* revision history
   hm  10. dec 2007  rev 1.0
     original version

   hm  17. sep. 2007 rev 1.1
     improved performance

   hm  21. jul. 2009 rev 1.2
     fixed a timing probelm


   *)
END_FUNCTION_BLOCK

FUNCTION_BLOCK "TP_1"   // FB67, SCL
TITLE = TP_1
{ S7_Optimized_Access := 'FALSE' }
AUTHOR : hugo
FAMILY : GENERAT
NAME : TP_1
VERSION : 1.0
// TP_1 generates a pulse every time it is calles with in := TRUE.
// in addition the timer can be cleared asynchronously with rst.
// the timer can be retriggered as often as necessary. it will count PT from the last trigger.
// 
// uses: T_PLC_MS [FC64]
//       STIME [FB64],IDB_STIME [DB64]
   VAR_INPUT
      IN : Bool;
      PT : Time;
      RST : Bool;
   END_VAR
   VAR_OUTPUT
      Q : Bool;
   END_VAR
   VAR
      tx : Time;
      start : Time;
      ix : Bool;
   END_VAR
BEGIN


   (* read system timer *)
   #tx := T_CONV(DWORD_TO_DINT("T_PLC_MS"()));

   IF #RST THEN
       #Q := FALSE;
   ELSIF #IN AND NOT #ix THEN
       #Q := TRUE;
       #start := #tx;
   ELSIF #tx - #start >= #PT THEN
       #Q := FALSE;
   END_IF;

   #ix:= #IN;



   (* revision history
   hm  28. jun. 2008
       original version

   *)
END_FUNCTION_BLOCK

FUNCTION_BLOCK "TP_1D"   // FB68, SCL
TITLE = TP_1D
{ S7_Optimized_Access := 'FALSE' }
AUTHOR : hugo
FAMILY : GENERAT
NAME : TP_1D
VERSION : 1.0
// TP_2 generates a pulse every time it is calles with in := TRUE.
// the module will reset IN by itself so no clearing of in is necessary.
// in addition the timer can be cleared asynchronously with rst.
// also the rst input is cleared by the module itself.
// the timer can be retriggered as often as necessary. it will count PT from the last trigger.
// after the time PT1 is elapsed, the timer blocks itself for PT2 and only allow new sequences after PT2 has elapsed.
// 
// uses: T_PLC_MS [FC64]
//       STIME [FB64],IDB_STIME [DB64]
   VAR_INPUT
      IN : Bool;
      PT1 : Time;
      PTD : Time;
      RST : Bool;
   END_VAR
   VAR_OUTPUT
      Q : Bool;
      W : Bool;
   END_VAR
   VAR
      tx : Time;
      start : Time;
      ix : Bool;
   END_VAR
BEGIN


   (* read system timer *)
   #tx := T_CONV(DWORD_TO_DINT("T_PLC_MS"()));

   IF #RST THEN
       #Q := FALSE;
       #RST := FALSE;
       #W := FALSE;
   ELSIF #W THEN
       IF #tx - #start >= #PTD THEN
           #W := FALSE;
       END_IF;
   ELSIF #IN AND NOT #ix THEN
       #Q := TRUE;
       #start := #tx;
       #IN := FALSE;
   ELSIF #tx - #start >= #PT1 THEN
       #Q := FALSE;
       #W := TRUE;
       #start := #tx;
   END_IF;

   #ix := #IN;



   (* revision history
   hm  28. jun. 2008
       original version

   *)
END_FUNCTION_BLOCK

FUNCTION_BLOCK "TP_X"   // FB69, SCL
TITLE = TP_X
{ S7_Optimized_Access := 'FALSE' }
AUTHOR : hugo
FAMILY : GENERAT
NAME : TP_R
VERSION : 1.3
// retriggerable edge triggered pulse similar to TP but with a retrigger function
// if the pt input is 0 then output is always low.
// 
// uses: T_PLC_MS [FC64]
//       STIME [FB64],IDB_STIME [DB64]
   VAR_INPUT
      IN : Bool;
      PT : Time;
   END_VAR
   VAR_OUTPUT
      Q : Bool;
      ET : Time;
   END_VAR
   VAR
      edge : Bool;
      start : Time;
      tx : Time;
   END_VAR
   VAR_TEMP
      TOP_SI : Struct
         EV_CLASS : Byte;
         EV_NUM : Byte;
         PRIORITY : Byte;
         NUM : Byte;
         TYP2_3 : Byte;
         TYP1 : Byte;
         ZI1 : Word;
         ZI2_3 : DWord;
      END_STRUCT;
      START_UP_SI : Struct
         EV_CLASS : Byte;
         EV_NUM : Byte;
         PRIORITY : Byte;
         NUM : Byte;
         TYP2_3 : Byte;
         TYP1 : Byte;
         ZI1 : Word;
         ZI2_3 : DWord;
      END_STRUCT;
      ERR : Int;
   END_VAR
BEGIN


   (* read actual startup info *)
   (* OB1_SCAN_1  BYTE  -  B#16#01: Abschluss des Neustarts (Warmstarts)
                        -  B#16#02: Abschluss des Wiederanlaufs
                        -  B#16#03: Abschluss des freien Zyklus
                        -  B#16#04: Abschluss des Kaltstarts
                        -  B#16#05: Erster OB 1-Zyklus der neuen Master-CPU nach 
                                    Master-Reserve-Umschaltung und STOP des 
                                    bisherigen Masters *)

   #ERR := RD_SINFO (TOP_SI => #TOP_SI, START_UP_SI => #START_UP_SI);

   (* read system_time *)
   #tx := T_CONV(DWORD_TO_DINT("T_PLC_MS"()));

   (* reset last_time on system startup *)
   IF #TOP_SI.EV_NUM = 1 OR #TOP_SI.EV_NUM = 2 OR #TOP_SI.EV_NUM = 4 THEN 
       #start := #tx;
   END_IF;

   (* rising edge trigger *)
   IF #IN AND NOT #edge THEN
       #start := #tx;
       #Q := #PT > t#0ms;
   ELSIF #Q THEN
       #ET := #tx - #start;
       IF #ET >= #PT THEN
           #Q := FALSE;
           #ET := t#0ms;
       END_IF;
   END_IF;
   #edge := #IN;


   (* revision history
   hm  4. aug 2006     rev 1.0
       original version

   hm  17. sep 2007    rev 1.1
       replaced time() with T_PLC_MS() for compatibility reasons

   hm  19. oct. 2008   rev 1.2
       renamed to TP_R to TP_X for compatibility reasons

   hm  17. dec. 2008   rev 1.3
       code optimized

   *)
END_FUNCTION_BLOCK

FUNCTION_BLOCK "CYCLE_4"   // FB239, SCL
TITLE = CYCLE_4
{ S7_Optimized_Access := 'FALSE' }
AUTHOR : hugo
FAMILY : GENERAT
NAME : CYCLE4
VERSION : 1.0
// uses: T_PLC_MS [FC64]
//       STIME [FB64],IDB_STIME [DB64]
   VAR_INPUT
      "E" : Bool := TRUE;
      T0 : Time;
      T1 : Time;
      T2 : Time;
      T3 : Time;
      S0 : Bool;
      SX : Int;
      SL : Bool;
   END_VAR
   VAR_OUTPUT
      STATE : Int;
   END_VAR
   VAR
      tx : Time;
      last : Time;
      init : Bool;
   END_VAR
   VAR_TEMP
      TOP_SI : Struct
         EV_CLASS : Byte;
         EV_NUM : Byte;
         PRIORITY : Byte;
         NUM : Byte;
         TYP2_3 : Byte;
         TYP1 : Byte;
         ZI1 : Word;
         ZI2_3 : DWord;
      END_STRUCT;
      START_UP_SI : Struct
         EV_CLASS : Byte;
         EV_NUM : Byte;
         PRIORITY : Byte;
         NUM : Byte;
         TYP2_3 : Byte;
         TYP1 : Byte;
         ZI1 : Word;
         ZI2_3 : DWord;
      END_STRUCT;
      ERR : Int;
   END_VAR
BEGIN


   (* read actual startup info *)
   (* OB1_SCAN_1  BYTE  -  B#16#01: Abschluss des Neustarts (Warmstarts)
                        -  B#16#02: Abschluss des Wiederanlaufs
                        -  B#16#03: Abschluss des freien Zyklus
                        -  B#16#04: Abschluss des Kaltstarts
                        -  B#16#05: Erster OB 1-Zyklus der neuen Master-CPU nach 
                                    Master-Reserve-Umschaltung und STOP des 
                                    bisherigen Masters *)

     #ERR := RD_SINFO (TOP_SI => #TOP_SI, START_UP_SI => #START_UP_SI);

   (* reset last_time on system startup *)
   IF #TOP_SI.EV_NUM = 1 OR #TOP_SI.EV_NUM = 2 OR #TOP_SI.EV_NUM = 4 THEN 
       #init := false;
   END_IF;

   (* read system timer *)
   #tx := T_CONV(DWORD_TO_DINT("T_PLC_MS"()));
   (* init on first cycle *)
   IF NOT #init THEN
       #init := TRUE;
       #last := #tx;
   END_IF;

   IF #"E" THEN
       IF #SL THEN
           (* when sx > 0 then the state sx is forced to start *)
           #STATE:= LIMIT(MN:=0,IN:=#SX,MX:=3);
           #last := #tx;
           (* this is to avoid to reset sx from the calling programm it does work fine on codesys but i am not sure about other systems, because we are writing to an input *)
           #SL := FALSE;
       ELSE
           CASE #STATE OF
               0 : (* wait for T0 and switch to next cycle *)
                   IF #tx - #last >= #T0 THEN
                       #STATE := 1;
                       #last := #tx;
                   END_IF;
               1 : (* wait for T1 over 1st cycle *)
                   IF #tx - #last >= #T1 THEN
                       #STATE := 2;
                       #last := #tx;
                   END_IF;
               2 : (* wait for T1 over 1st cycle *)
                   IF #tx - #last >= #T2 THEN
                       #STATE := 3;
                       #last := #tx;
                   END_IF;
               3 : (* wait for T2 over 2nd cycle *)
                   IF #tx - #last >= #T3 THEN
                       IF #S0 THEN #STATE := 0; END_IF; (* if S0 is false, the sequence stops at state 3 *)
                       #last := #tx;
                   END_IF;
           END_CASE;
       END_IF;
   ELSE
       #STATE := 0;
       #last := #tx;
   END_IF;


   (*
   hm  3. nov. 2008 rev 1.0
       original version

   *)
END_FUNCTION_BLOCK

FUNCTION "T_PLC_MS" : DWord   // FC64, SCL
TITLE = T_PLC_MS
{ S7_Optimized_Access := 'FALSE' }
AUTHOR : hugo
FAMILY : MEASURE
NAME : T_PLC_MS
VERSION : 1.2
// T_PLC_MS reads the internal PLC timer and return the time, it has the advantage to be able to set a debug mode 
// and speed up the counter to test the plc timer overrun which occurs every 50 days respectively 25 days at siemens S7
// this routine also allows to correct the behavior of s7 where the internal plc counter will not count all 32 bits.
// 
// uses: STIME [FB64],IDB_STIME [DB64]
BEGIN


   "IDB_STIME"(); 
   #T_PLC_MS := "IDB_STIME".tx; 
   (* hier muss die korrektur für step7 stattfinden
   plctime muss den vollen wertebereich von time ausnutzen:
   wenn bei step7 time -24tage bis plus 24 tage ist dann muss der timer auch beim überlauf auf -24tage springen 
   und auf keinen fall auf 0 !!!!
   für siemens muss ein weiterer fb im main eingebunden werden der sicherstellt das alle 32 bits durchgezählt werden.
   es kann nur ein fb sein den er muss sich das oberste (32te) bit merken.
   oder etwa spring s7 bei überlauf auf -24 tage????? dann wäre keine korrektur nötig.
   *)
   IF "debug" THEN
       #T_PLC_MS := DINT_TO_DWORD((DWORD_TO_DINT(SHL(IN:=#T_PLC_MS,N:="N") OR SHL(IN:=DWORD#1,N:="N"))-1) + DWORD_TO_DINT("offset_1"));
   END_IF;


   (* revision history
   hm  14.9.2007   rev 1.0
       original version

   hm  12. nov 2007    rev 1.1
       added temporaray variable tx because some compilers could not handle time() as an argument

   hm  16. nov. 2008   rev 1.2
       initialized constants with 0 for compatibility reasons
   *)
END_FUNCTION

FUNCTION "INC2" : Int   // FC91, SCL
TITLE = INC2
{ S7_Optimized_Access := 'FALSE' }
AUTHOR : hugo
FAMILY : MATH
NAME : INC2
VERSION : 1.0
// This function increments the input X by the value D and compares the result with U.
// if the output exceeds U it will continue to count from L again.
   VAR_INPUT
      X : Int;
      D : Int;
      L : Int;
      U : Int;
   END_VAR
   VAR_TEMP
      tmp : Int;
   END_VAR
BEGIN


   #tmp := #U - #L + 1;
   #INC2 := (#X + #D - #L + #tmp) MOD #tmp + #L;



   (* revision history
   hm  29. jun. 2008       REV 1.0
       original version


   *)
END_FUNCTION

// ===== PLC "Logic memory"  Unspecific CPU S7 300 =====

VAR_GLOBAL CONSTANT   // PLC tag table "STEP7 classic symbols"
   "n" : Int := 16;
   "n_FB38" : Int := 32;   // MigChange: n
   "N(1)" : Int := 15;
   "n_FB40" : Int := 31;   // MigChange: n
END_VAR

FUNCTION_BLOCK "FIFO_16"   // FB37, SCL
TITLE = FIFO_16
{ S7_Optimized_Access := 'FALSE' }
AUTHOR : hugo
FAMILY : MEMORY
NAME : FIFO_16
VERSION : 2.0
// 16 Dword FIFO memory
// 
// uses: INC1 [FC53]
   VAR_INPUT
      Din : DWord;
      "E" : Bool := TRUE;
      RD : Bool;
      WD : Bool;
      RST : Bool;
   END_VAR
   VAR_OUTPUT
      Dout : DWord;
      EMPTY : Bool := TRUE;
      FULL : Bool;
   END_VAR
   VAR
      fifo : Array[0..16] of DWord;
      pr : Int;
      pw : Int;
   END_VAR
BEGIN


   IF #RST THEN
     #pw := #pr;
     #FULL := FALSE;
     #EMPTY := TRUE;
     #Dout := 0;
   ELSIF #"E" THEN
     IF NOT #EMPTY AND #RD THEN
       #Dout := #fifo[#pr];
       #pr := "INC1"(X:=#pr,N:="n");
       #EMPTY := #pr = #pw;
       #FULL := FALSE;
     END_IF;
     IF NOT #FULL AND #WD THEN
       #fifo[#pw] := #Din;
       #pw := "INC1"(X:=#pw,N:="n");
       #FULL := #pw = #pr;
       #EMPTY := FALSE;
     END_IF;
   END_IF;


   (* revision history

   hm  4. aug. 2006  rev 1.0
     original version

   hm  19. feb 2008 rev 1.1
     performance improvements

   hm  17. oct. 2008 rev 1.2
     improved performance

   ks  27. oct. 2008 rev 1.3
     optimized coding

   hm  14. mar. 2009 rev 1.4
     removed double assignments

   hm 24. jul. 2009  rev 2.0
     chaged inputs E and WR to E, WD and WR
     allow read and write in one cycle

   *)
END_FUNCTION_BLOCK

FUNCTION_BLOCK "FIFO_32"   // FB38, SCL
TITLE = FIFO_32
{ S7_Optimized_Access := 'FALSE' }
AUTHOR : hugo
FAMILY : MEMORY
NAME : FIFO_32
VERSION : 2.0
// 32 Dword FIFO memory
// 
// uses: INC1 [FC53]
   VAR_INPUT
      Din : DWord;
      "E" : Bool := TRUE;
      RD : Bool;
      WD : Bool;
      RST : Bool;
   END_VAR
   VAR_OUTPUT
      Dout : DWord;
      EMPTY : Bool := TRUE;
      FULL : Bool;
   END_VAR
   VAR
      fifo : Array[0..32] of DWord;
      pr : Int;
      pw : Int;
   END_VAR
BEGIN


   IF #RST THEN
     #pw := #pr;
     #FULL := FALSE;
     #EMPTY := TRUE;
     #Dout := 0;
   ELSIF #"E" THEN
     IF NOT #EMPTY AND #RD THEN
       #Dout := #fifo[#pr];
       #pr := "INC1"(X:=#pr,N:="n_FB38");
       #EMPTY := #pr = #pw;
       #FULL := FALSE;
     END_IF;
     IF NOT #FULL AND #WD THEN
       #fifo[#pw] := #Din;
       #pw := "INC1"(X:=#pw,N:="n_FB38");
       #FULL := #pw = #pr;
       #EMPTY := FALSE;
     END_IF;
   END_IF;

   (* revision history
   hm  4. aug. 2006  rev 1.0
     original version

   hm  19. feb 2008  rev 1.1
     performance improvements

   hm  17. oct. 2008 rev 1.2
     improved performance

   ks  27. oct. 2008 rev 1.3
     improved code

   hm  14. mar. 2009 rev 1.4
     removed double assignments

   hm 24. jul. 2009  rev 2.0
     chaged inputs E and WR to E, WD and WR
     allow read and write in one cycle

   *)
END_FUNCTION_BLOCK

FUNCTION_BLOCK "STACK_16"   // FB39, SCL
TITLE = STACK_16
{ S7_Optimized_Access := 'FALSE' }
AUTHOR : hugo
FAMILY : MEMORY
NAME : STACK_16
VERSION : 2.0
// 16 Dword STACK memory
   VAR_INPUT
      Din : DWord;
      "E" : Bool := TRUE;
      RD : Bool;
      WD : Bool;
      RST : Bool;
   END_VAR
   VAR_OUTPUT
      Dout : DWord;
      EMPTY : Bool := TRUE;
      FULL : Bool;
   END_VAR
   VAR
      stack : Array[0..15] of DWord;
      pt : Int;
   END_VAR
BEGIN


   IF #RST THEN
     (* asynchronous reset for the fifo *)
     #pt := 0;
     #EMPTY := TRUE;
     #FULL := FALSE;
     #Dout := 0;
   ELSIF #"E" THEN
     IF NOT #EMPTY AND #RD THEN
       (* read one element *)
       #pt := #pt - 1;
       #Dout := #stack[#pt];
       #EMPTY := #pt = 0;
       #FULL := FALSE;
     END_IF;
     IF NOT #FULL AND #WD THEN
       (* write one element *)
       #stack[#pt] := #Din;
       #pt := #pt + 1;
       #FULL := #pt > "n";
       #EMPTY := FALSE;
     END_IF;
   END_IF;


   (* revision history
   hm  4. aug. 2006  rev 1.0
     original version

   hm  19. feb 2008  rev 1.1
     performance improvements

   hm  17. oct. 2008 rev 1.2
     deleted unnecessary init with 0

   hm  27. oct. 2008 rev 1.3
     optimized performance

   hm  25. jul 2009  rev 2.0
     changed inputs to allow simultsaneous read and write
   *)
END_FUNCTION_BLOCK

FUNCTION_BLOCK "STACK_32"   // FB40, SCL
TITLE = STACK_32
{ S7_Optimized_Access := 'FALSE' }
AUTHOR : hugo
FAMILY : MEMORY
NAME : STACK_32
VERSION : 2.0
// 32 Dword STACK memory
   VAR_INPUT
      Din : DWord;
      "E" : Bool := TRUE;
      RD : Bool;
      WD : Bool;
      RST : Bool;
   END_VAR
   VAR_OUTPUT
      Dout : DWord;
      EMPTY : Bool := TRUE;
      FULL : Bool;
   END_VAR
   VAR
      stack : Array[0..31] of DWord;
      pt : Int;
   END_VAR
BEGIN


   IF #RST THEN
     (* asynchronous reset for the fifo *)
     #pt := 0;
     #EMPTY := TRUE;
     #FULL := FALSE;
     #Dout := 0;
   ELSIF #"E" THEN
     IF NOT #EMPTY AND #RD THEN
       (* read one element *)
       #pt := #pt - 1;
       #Dout := #stack[#pt];
       #EMPTY := #pt = 0;
       #FULL := FALSE;
     END_IF;
     IF NOT #FULL AND #WD THEN
       (* write one element *)
       #stack[#pt] := #Din;
       #pt := #pt + 1;
       #FULL := #pt > "n_FB40";
       #EMPTY := FALSE;
     END_IF;
   END_IF;


   (* revision history
   hm  4. aug. 2006  rev 1.0
     original version

   hm  19. feb 2008  rev 1.1
     performance improvements

   hm  17. oct. 2008 rev 1.2
     deleted unnecessary init with 0

   ks  27. oct. 2008 rev 1.3
     optimized performance

   hm  25. jul 2009  rev 2.0
     changed inputs to allow simultsaneous read and write

   *)
END_FUNCTION_BLOCK

FUNCTION "INC1" : Int   // FC53, SCL
TITLE = INC1
{ S7_Optimized_Access := 'FALSE' }
AUTHOR : hugo
FAMILY : MATH
NAME : INC1
VERSION : 1.2
// This is a increment function which increments the variable X by 1 and if M is reached, it begins with 0 again.
// _inc1(3,X) will generate 0,1,2,3,0,1,.....
   VAR_INPUT
      X : Int;
      N : Int;
   END_VAR
BEGIN


   IF #X >= #N - 1 THEN
       #INC1 := 0;
   ELSE
       #INC1 := #X + 1;
   END_IF;


   (* this elegant version is 50% slower
   INC1 := X := (x + 1) MOD N;
   *)



   (* revision history
   hm  13. oct. 2008   rev 1.0
       original version

   hm  22. oct. 2008   rev 1.1
       added statement to return value for compatibility reasons

   hm  23. feb. 2009   rev 1.2
       when inc1 is called with X >= N inc will continue with 0
   *)
END_FUNCTION

// ===== PLC "Math Double Precision"  Unspecific CPU S7 300 =====

TYPE "REAL2"
VERSION : 0.0
   STRUCT
      R1 : Real;
      RX : Real;
   END_STRUCT;
END_TYPE

FUNCTION "R2_ABS" : "REAL2"   // FC143, SCL
TITLE = R2_ABS
{ S7_Optimized_Access := 'FALSE' }
AUTHOR : hugo
FAMILY : R2
NAME : ABS
VERSION : 1.1
// R2_abs returns the absulute value of a double precision real.
//  
// uses: REAL2 [UDT11]
   VAR_INPUT
      X : "REAL2";
   END_VAR
   VAR_TEMP
      tR2_ABS : "REAL2";
   END_VAR
BEGIN


   IF #X.RX >= 0.0 THEN
       #tR2_ABS.RX := #X.RX;
       #tR2_ABS.R1 := #X.R1;
   ELSE
       #tR2_ABS.RX := -#X.RX;
       #tR2_ABS.R1 := -#X.R1;
   END_IF;

   #R2_ABS := #tR2_ABS;


